screen "MTA-CompALTA" 1280x800, template "Plantilla"
   GraphicIOField "Plantilla_Campo ES gráfico_3" at 758,425 size 65x60
   GraphicIOField "Plantilla_Campo ES gráfico_4" at 685,353 size 65x60
   GraphicIOField "Plantilla_Campo ES gráfico_5" at 612,281 size 65x60
   GraphicIOField "Plantilla_Campo ES gráfico_2" at 539,209 size 65x60
   GraphicView "Visor de gráficos_2" at 492,46 size 254x172
   GraphicView "Visor de gráficos_18" at 492,46 size 254x172
   GraphicIOField "Plantilla_Campo ES gráfico_1" at 490,113 size 100x102
   GraphicView "Visor de gráficos_3" at 569,134 size 246x148
   ScreenModuleView "Faceplate_8_1" at 781,145 size 47x30
   GraphicView "Visor de gráficos_8" at 1175,577 size 29x50
   GraphicView "Visor de gráficos_7" at 885,605 size 391x113
   TextField "Plantilla_Campo de texto_1" at 1141,578 size 32x23
   IOField "Campo ES_1" at 943,632 size 108x28
   Button "Botón_7" at 1119,186 size 128x41
   Button "Botón_12" at 1119,234 size 128x41
   Button "Botón_13" at 1119,138 size 128x41
   Button "Botón_14" at 641,627 size 160x46
   TextField "Campo de texto_2" at 519,9 size 242x27
   ScreenModuleView "Faceplate_8_5" at 927,289 size 47x30
   ScreenModuleView "Faceplate_8_4" at 1000,361 size 47x30
   GraphicView "Visor de gráficos_19" at 569,134 size 246x148
   ScreenModuleView "Faceplate_8_2" at 854,217 size 47x30
   GraphicView "Visor de gráficos_4" at 642,206 size 246x148
   GraphicView "Visor de gráficos_22" at 642,206 size 246x148
   GraphicView "Visor de gráficos_5" at 715,278 size 246x148
   GraphicView "Visor de gráficos_21" at 715,278 size 246x148
   GraphicView "Visor de gráficos_6" at 788,350 size 246x148
   GraphicView "Visor de gráficos_20" at 788,350 size 246x148
   ScreenModuleView "Faceplate_8_3" at 1072,433 size 47x30
   ScreenModuleView "Faceplate_8_6" at 748,113 size 47x30
   Button "Botón_3" at 1181,68 size 48x46
   ScreenModuleView "Faceplate_8_7" at 1144,505 size 47x30
   GraphicIOField "Plantilla_Campo ES gráfico_6" at 831,497 size 65x60
   GraphicView "Visor de gráficos_1" at 861,422 size 246x148
   GraphicView "Visor de gráficos_9" at 861,422 size 246x148
   GraphicIOField "Campo ES gráfico_4" at 6,182 size 374x6
   SymbolicIOField "Campo ES simbólico_4" at 25,154 size 178x21
   TextField "Campo de texto_1" at 19,121 size 55x32
   GraphicIOField "Campo ES gráfico_5" at 118,341 size 374x6
   TextField "Campo de texto_6" at 127,280 size 67x32
   SymbolicIOField "Campo ES simbólico_5" at 137,313 size 186x21
   GraphicIOField "Campo ES gráfico_1" at 191,422 size 374x6
   TextField "Campo de texto_8" at 200,361 size 67x32
   SymbolicIOField "Campo ES simbólico_1" at 210,394 size 186x21
   GraphicIOField "Campo ES gráfico_3" at 44,262 size 373x6
   TextField "Campo de texto_10" at 53,201 size 67x32
   SymbolicIOField "Campo ES simbólico_3" at 63,234 size 194x21
   GraphicIOField "Campo ES gráfico_2" at 264,502 size 374x6
   TextField "Campo de texto_9" at 273,441 size 67x32
   SymbolicIOField "Campo ES simbólico_2" at 283,474 size 186x21
   GraphicIOField "Campo ES gráfico_16" at 337,582 size 374x6
   TextField "Campo de texto_3" at 346,521 size 67x32
   SymbolicIOField "Campo ES simbólico_11" at 356,554 size 186x21
   IOField "Campo ES_6" at 255,157 size 85x19
   IOField "Campo ES_2" at 367,316 size 85x19
   IOField "Campo ES_3" at 439,397 size 85x19
   IOField "Campo ES_5" at 292,237 size 85x19
   IOField "Campo ES_4" at 512,477 size 85x19
   IOField "Campo ES_7" at 585,557 size 85x19
   ScreenModuleView "Faceplate_6_1" at 283,125 size 57x28
   ScreenModuleView "Faceplate_6_5" at 395,284 size 57x28
   ScreenModuleView "Faceplate_6_4" at 468,365 size 57x28
   ScreenModuleView "Faceplate_6_2" at 321,205 size 57x28
   ScreenModuleView "Faceplate_6_3" at 541,445 size 57x28
   GraphicIOField "Campo ES gráfico_6" at 348,125 size 9x45
   GraphicIOField "Campo ES gráfico_9" at 357,125 size 9x45
   SymbolicIOField "Campo ES simbólico_6" at 86,124 size 160x29
   Button "Botón_11" at 6,116 size 374x64
   Switch "Interruptor_1" at 250,125 size 29x29
   Switch "Interruptor_10" at 863,114 size 40x40
   GraphicIOField "Campo ES gráfico_14" at 459,286 size 9x45
   GraphicIOField "Campo ES gráfico_15" at 468,286 size 9x45
   SymbolicIOField "Campo ES simbólico_10" at 195,283 size 160x29
   Button "Botón_6" at 118,275 size 374x64
   Switch "Interruptor_5" at 360,285 size 29x29
   Switch "Interruptor_9" at 1009,258 size 40x40
   GraphicIOField "Campo ES gráfico_12" at 532,367 size 9x45
   GraphicIOField "Campo ES gráfico_13" at 541,367 size 9x45
   Button "Botón_8" at 191,356 size 374x64
   SymbolicIOField "Campo ES simbólico_9" at 269,364 size 160x29
   Switch "Interruptor_4" at 433,366 size 29x29
   Switch "Interruptor_8" at 1082,330 size 40x40
   GraphicIOField "Campo ES gráfico_7" at 385,207 size 9x45
   GraphicIOField "Campo ES gráfico_10" at 394,207 size 9x45
   SymbolicIOField "Campo ES simbólico_7" at 120,204 size 160x29
   Switch "Interruptor_6" at 936,186 size 40x40
   GraphicIOField "Campo ES gráfico_8" at 605,447 size 9x45
   GraphicIOField "Campo ES gráfico_11" at 614,447 size 9x45
   SymbolicIOField "Campo ES simbólico_8" at 341,444 size 160x29
   Button "Botón_9" at 264,436 size 374x64
   Switch "Interruptor_3" at 504,445 size 29x29
   Switch "Interruptor_7" at 1155,402 size 40x40
   Switch "Interruptor_11" at 1228,474 size 40x40
   ScreenModuleView "Faceplate_6_6" at 614,525 size 57x28
   GraphicIOField "Campo ES gráfico_17" at 678,527 size 9x45
   GraphicIOField "Campo ES gráfico_18" at 687,527 size 9x45
   SymbolicIOField "Campo ES simbólico_12" at 414,524 size 160x29
   Button "Botón_1" at 337,516 size 374x64
   Switch "Interruptor_12" at 577,525 size 29x29
   Button "Botón_10" at 45,196 size 374x64
   Switch "Interruptor_2" at 284,206 size 29x29
   TextField "Campo de texto_4" at 591,208 size 309x29
   Button "Botón_2" at 912,202 size 128x41

screen "MTA-ALTAMC006" 1280x800, template "Plantilla-Alta-Cmp"
   Button "Botón_1" at 186,441 size 48x38
   Button "Botón_2" at 186,401 size 48x38
   Button "Botón_7" at 390,106 size 40x38
   Button "Botón_8" at 306,600 size 96x35
   TextField "Campo de texto_6" at 266,362 size 72x27
   TextField "Campo de texto_7" at 82,426 size 84x27
   TextField "Campo de texto_8" at 362,363 size 40x27
   TextField "Campo de texto_11" at 26,343 size 158x27
   GraphicIOField "Campo ES gráfico_3" at 294,402 size 16x78
   GraphicIOField "Campo ES gráfico_5" at 374,402 size 16x78
   SymbolicIOField "Campo ES simbólico_2" at 9,290 size 424x37
   TextField "Campo de texto_16" at 521,10 size 279x27
   TextField "Campo de texto_1" at 32,510 size 326x27
   TextField "Campo de texto_4" at 32,570 size 231x27
   TextField "Campo de texto_5" at 32,635 size 231x27
   Button "Botón_3" at 306,665 size 96x35
   GraphicIOField "Campo ES gráfico_2" at 10,280 size 422x6
   SymbolicIOField "Campo ES simbólico_4" at 19,246 size 290x21
   Button "Botón_6" at 13,154 size 88x62
   Switch "Interruptor_1" at 150,167 size 37x37
   ScreenModuleView "Faceplate_6_1" at 342,236 size 76x34
   ScreenModuleView "Faceplate_7_1" at 213,158 size 207x70
   IOField "Campo ES_7" at 20,535 size 173x35
   IOField "Campo ES_1" at 200,535 size 80x35
   IOField "Campo ES_2" at 20,595 size 173x35
   IOField "Campo ES_3" at 20,660 size 173x35

screen "EPROC-ALTAMS050" 1280x800, template "Plantilla-Alta-Sec"
   Button "Botón_3" at 467,294 size 40x38
   Button "Botón_4" at 411,540 size 96x35
   TextField "Campo de texto_6" at 37,450 size 326x27
   TextField "Campo de texto_4" at 37,510 size 201x27
   IOField "Campo ES_7" at 25,475 size 173x35
   IOField "Campo ES_1" at 205,475 size 80x35
   IOField "Campo ES_2" at 25,535 size 173x35
   GraphicIOField "Campo ES gráfico_3" at 21,434 size 511x6
   TextField "Campo de texto_3" at 46,356 size 89x39
   SymbolicIOField "Campo ES simbólico_3" at 48,392 size 242x21
   Switch "Interruptor_8" at 205,359 size 29x29
   ScreenModuleView "Faceplate_2_4" at 274,346 size 244x69

screen "EPROC-ALTAMS051" 1280x800, template "Plantilla-Alta-Sec"
   Button "Botón_3" at 467,294 size 40x38
   Button "Botón_4" at 411,540 size 96x35
   TextField "Campo de texto_6" at 37,450 size 326x27
   TextField "Campo de texto_4" at 37,510 size 201x27
   IOField "Campo ES_7" at 25,475 size 173x35
   IOField "Campo ES_1" at 205,475 size 80x35
   IOField "Campo ES_2" at 25,535 size 173x35
   GraphicIOField "Campo ES gráfico_9" at 21,434 size 511x6
   TextField "Campo de texto_1" at 46,356 size 89x39
   SymbolicIOField "Campo ES simbólico_9" at 48,392 size 242x21
   Switch "Interruptor_5" at 211,363 size 29x29
   ScreenModuleView "Faceplate_2_1" at 277,346 size 244x69

screen "EPROC-ALTAMS052" 1280x800, template "Plantilla-Alta-Sec"
   Button "Botón_3" at 467,294 size 40x38
   Button "Botón_4" at 411,540 size 96x35
   TextField "Campo de texto_6" at 37,450 size 326x27
   TextField "Campo de texto_4" at 37,510 size 201x27
   IOField "Campo ES_7" at 25,475 size 173x35
   IOField "Campo ES_1" at 205,475 size 80x35
   IOField "Campo ES_2" at 25,535 size 173x35
   GraphicIOField "Campo ES gráfico_1" at 21,434 size 511x6
   TextField "Campo de texto_1" at 46,356 size 89x39
   SymbolicIOField "Campo ES simbólico_1" at 48,392 size 242x21
   Switch "Interruptor_6" at 227,365 size 29x29
   ScreenModuleView "Faceplate_2_2" at 277,346 size 244x69

screen "EPROC-ALTAMS053" 1280x800, template "Plantilla-Alta-Sec"
   Button "Botón_3" at 467,294 size 40x38
   Button "Botón_4" at 411,540 size 96x35
   TextField "Campo de texto_6" at 37,450 size 326x27
   TextField "Campo de texto_4" at 37,510 size 201x27
   IOField "Campo ES_7" at 25,475 size 173x35
   IOField "Campo ES_1" at 205,475 size 80x35
   IOField "Campo ES_2" at 25,535 size 173x35
   IOField "Campo ES_6" at 351,413 size 85x19
   GraphicIOField "Campo ES gráfico_2" at 21,434 size 511x6
   TextField "Campo de texto_2" at 46,351 size 101x39
   SymbolicIOField "Campo ES simbólico_2" at 48,387 size 242x21
   Switch "Interruptor_7" at 227,360 size 29x29
   ScreenModuleView "Faceplate_2_3" at 276,346 size 244x69

screen "EPROC-BAJAMC060" 1280x800, template "Plantilla-Baja-Cmp"
   Button "Botón_4" at 1135,405 size 96x35
   TextField "Campo de texto_6" at 761,315 size 326x27
   TextField "Campo de texto_4" at 761,375 size 231x27
   Button "Botón_1" at 1135,470 size 96x35
   TextField "Campo de texto_1" at 761,440 size 231x27
   Button "Botón_2" at 1135,535 size 96x35
   TextField "Campo de texto_2" at 761,505 size 231x27
   Button "Botón_3" at 1135,600 size 96x35
   TextField "Campo de texto_3" at 761,570 size 231x27
   Button "Botón_5" at 1135,665 size 96x35
   TextField "Campo de texto_7" at 761,635 size 231x27
   Button "Botón_6" at 1199,168 size 40x38
   GraphicIOField "Campo ES gráfico_4" at 746,294 size 511x6
   TextField "Campo de texto_5" at 771,224 size 116x39
   SymbolicIOField "Campo ES simbólico_9" at 773,260 size 242x21
   Switch "Interruptor_5" at 1108,242 size 91x31
   IOField "Campo ES_7" at 749,340 size 173x35
   IOField "Campo ES_1" at 929,340 size 80x35
   IOField "Campo ES_2" at 749,400 size 173x35
   IOField "Campo ES_3" at 749,465 size 173x35
   IOField "Campo ES_4" at 749,530 size 173x35
   IOField "Campo ES_5" at 749,595 size 173x35
   IOField "Campo ES_6" at 749,660 size 173x35

screen "EPROC-BAJAMC061" 1280x800, template "Plantilla-Baja-Cmp"
   Button "Botón_4" at 1135,405 size 96x35
   TextField "Campo de texto_6" at 761,315 size 326x27
   TextField "Campo de texto_4" at 761,375 size 231x27
   Button "Botón_1" at 1135,470 size 96x35
   TextField "Campo de texto_1" at 761,440 size 231x27
   Button "Botón_2" at 1135,535 size 96x35
   TextField "Campo de texto_2" at 761,505 size 231x27
   Button "Botón_3" at 1135,600 size 96x35
   TextField "Campo de texto_3" at 761,570 size 231x27
   Button "Botón_5" at 1135,665 size 96x35
   TextField "Campo de texto_7" at 761,635 size 231x27
   Button "Botón_6" at 1199,168 size 40x38
   IOField "Campo ES_7" at 749,340 size 173x35
   IOField "Campo ES_1" at 929,340 size 80x35
   IOField "Campo ES_2" at 749,400 size 173x35
   IOField "Campo ES_3" at 749,465 size 173x35
   IOField "Campo ES_4" at 749,530 size 173x35
   IOField "Campo ES_5" at 749,595 size 173x35
   IOField "Campo ES_6" at 749,660 size 173x35
   GraphicIOField "Campo ES gráfico_3" at 746,293 size 510x6
   TextField "Campo de texto_5" at 771,224 size 116x39
   SymbolicIOField "Campo ES simbólico_8" at 773,260 size 242x21
   Switch "Interruptor_4" at 974,228 size 29x29
   ScreenModuleView "Faceplate_1_1" at 1018,228 size 236x58

screen "EPROC-BAJAMC062" 1280x800, template "Plantilla-Baja-Cmp"
   Button "Botón_4" at 1135,405 size 96x35
   TextField "Campo de texto_6" at 761,315 size 326x27
   TextField "Campo de texto_4" at 761,375 size 231x27
   Button "Botón_1" at 1135,470 size 96x35
   TextField "Campo de texto_1" at 761,440 size 231x27
   Button "Botón_2" at 1135,535 size 96x35
   TextField "Campo de texto_2" at 761,505 size 231x27
   Button "Botón_3" at 1135,600 size 96x35
   TextField "Campo de texto_3" at 761,570 size 231x27
   Button "Botón_5" at 1135,665 size 96x35
   TextField "Campo de texto_7" at 761,635 size 231x27
   Button "Botón_6" at 1199,168 size 40x38
   IOField "Campo ES_7" at 749,340 size 173x35
   IOField "Campo ES_1" at 929,340 size 80x35
   IOField "Campo ES_2" at 749,400 size 173x35
   IOField "Campo ES_3" at 749,465 size 173x35
   IOField "Campo ES_4" at 749,530 size 173x35
   IOField "Campo ES_5" at 749,595 size 173x35
   IOField "Campo ES_6" at 749,660 size 173x35
   GraphicIOField "Campo ES gráfico_2" at 747,293 size 507x6
   TextField "Campo de texto_5" at 771,224 size 116x39
   SymbolicIOField "Campo ES simbólico_7" at 773,260 size 242x21
   Switch "Interruptor_3" at 970,227 size 29x29
   ScreenModuleView "Faceplate_1_3" at 1013,227 size 236x58

screen "EPROC-BAJAMC063" 1280x800, template "Plantilla-Baja-Cmp"
   Button "Botón_4" at 1135,405 size 96x35
   TextField "Campo de texto_6" at 761,315 size 326x27
   TextField "Campo de texto_4" at 761,375 size 231x27
   Button "Botón_1" at 1135,470 size 96x35
   TextField "Campo de texto_1" at 761,440 size 231x27
   Button "Botón_2" at 1135,535 size 96x35
   TextField "Campo de texto_2" at 761,505 size 231x27
   Button "Botón_3" at 1135,600 size 96x35
   TextField "Campo de texto_3" at 761,570 size 231x27
   Button "Botón_5" at 1135,665 size 96x35
   TextField "Campo de texto_7" at 761,635 size 231x27
   Button "Botón_6" at 1199,168 size 40x38
   IOField "Campo ES_7" at 749,340 size 173x35
   IOField "Campo ES_1" at 929,340 size 80x35
   IOField "Campo ES_2" at 749,400 size 173x35
   IOField "Campo ES_3" at 749,465 size 173x35
   IOField "Campo ES_4" at 749,530 size 173x35
   IOField "Campo ES_5" at 749,595 size 173x35
   IOField "Campo ES_6" at 749,660 size 173x35
   GraphicIOField "Campo ES gráfico_1" at 746,293 size 507x6
   TextField "Campo de texto_8" at 763,224 size 91x39
   SymbolicIOField "Campo ES simbólico_6" at 765,260 size 242x21
   Switch "Interruptor_2" at 967,227 size 29x29
   ScreenModuleView "Faceplate_1_4" at 1014,226 size 236x58

screen "EPROC-BAJAMC064" 1280x800, template "Plantilla-Baja-Cmp"
   Button "Botón_4" at 1135,405 size 96x35
   TextField "Campo de texto_6" at 761,315 size 326x27
   TextField "Campo de texto_4" at 761,375 size 231x27
   Button "Botón_1" at 1135,470 size 96x35
   TextField "Campo de texto_1" at 761,440 size 231x27
   Button "Botón_2" at 1135,535 size 96x35
   TextField "Campo de texto_2" at 761,505 size 231x27
   Button "Botón_3" at 1135,600 size 96x35
   TextField "Campo de texto_3" at 761,570 size 231x27
   Button "Botón_5" at 1135,665 size 96x35
   TextField "Campo de texto_7" at 761,635 size 231x27
   Button "Botón_6" at 1199,168 size 40x38
   IOField "Campo ES_7" at 749,340 size 173x35
   IOField "Campo ES_1" at 929,340 size 80x35
   IOField "Campo ES_2" at 749,400 size 173x35
   IOField "Campo ES_3" at 749,465 size 173x35
   IOField "Campo ES_4" at 749,530 size 173x35
   IOField "Campo ES_5" at 749,595 size 173x35
   IOField "Campo ES_6" at 749,660 size 173x35
   GraphicIOField "Campo ES gráfico_5" at 747,294 size 507x6
   TextField "Campo de texto_9" at 771,224 size 100x39
   SymbolicIOField "Campo ES simbólico_5" at 773,260 size 242x21
   Switch "Interruptor_1" at 969,227 size 29x29
   ScreenModuleView "Faceplate_1_5" at 1016,227 size 236x58

screen "EPROC-BAJAMS054" 1280x800, template "Plantilla-Baja-Sec"
   TextField "Campo de texto_1" at 758,509 size 326x27
   Button "Botón_4" at 1032,599 size 96x35
   TextField "Campo de texto_4" at 758,569 size 231x27
   TextField "Campo de texto_5" at 758,634 size 231x27
   Button "Botón_5" at 1032,664 size 96x35
   Button "Botón_6" at 1188,358 size 40x38
   IOField "Campo ES_7" at 746,534 size 173x35
   IOField "Campo ES_1" at 926,534 size 80x35
   IOField "Campo ES_2" at 746,594 size 173x35
   IOField "Campo ES_3" at 746,659 size 173x35
   GraphicIOField "Campo ES gráfico_3" at 736,489 size 510x6
   TextField "Campo de texto_6" at 761,411 size 116x39
   SymbolicIOField "Campo ES simbólico_8" at 763,447 size 242x21
   ScreenModuleView "Faceplate_3_1" at 1015,411 size 213x73

screen "EPROC-BAJAMS055" 1280x800, template "Plantilla-Baja-Sec"
   TextField "Campo de texto_1" at 758,509 size 326x27
   Button "Botón_4" at 1032,599 size 96x35
   TextField "Campo de texto_4" at 758,569 size 231x27
   TextField "Campo de texto_5" at 758,634 size 231x27
   Button "Botón_5" at 1032,664 size 96x35
   Button "Botón_6" at 1188,358 size 40x38
   IOField "Campo ES_7" at 746,534 size 173x35
   IOField "Campo ES_1" at 926,534 size 80x35
   IOField "Campo ES_2" at 746,594 size 173x35
   IOField "Campo ES_3" at 746,659 size 173x35
   GraphicIOField "Campo ES gráfico_4" at 736,489 size 511x6
   TextField "Campo de texto_2" at 761,411 size 116x39
   SymbolicIOField "Campo ES simbólico_9" at 763,447 size 242x21
   ScreenModuleView "Faceplate_3_2" at 1020,411 size 213x73

screen "Imagen_1" 1280x800
   GraphicIOField "Campo ES gráfico_3" at 736,489 size 510x6
   TextField "Campo de texto_6" at 761,411 size 116x39
   SymbolicIOField "Campo ES simbólico_8" at 763,447 size 242x21
   ScreenModuleView "Faceplate_3_1" at 1015,411 size 213x73

Template "Plantilla" 1280x800
   Button "Plantilla_6" at 1196,741 size 81x58
   Button "Plantilla_1" at 1037,749 size 78x50
   Button "Plantilla_3" at 717,748 size 78x50
   Button "Plantilla_4" at 877,748 size 78x50
   Button "Plantilla_5" at 957,748 size 78x50
   Button "Plantilla_7" at 479,748 size 78x50
   Button "Plantilla_8" at 161,748 size 78x50
   Button "Plantilla_9" at 81,748 size 78x50
   Button "Plantilla_10" at 1117,741 size 78x58
   Button "Plantilla_12" at 638,748 size 78x50
   Button "Plantilla_13" at 400,748 size 78x50
   Button "Plantilla_14" at 321,748 size 78x50
   Button "Plantilla_15" at 558,748 size 78x50
   Button "Plantilla_16" at 241,748 size 78x50
   Button "Plantilla_17" at 1,740 size 78x58
   GraphicView "Plantilla_Visor de gráficos_1" at 80,740 size 78x6
   GraphicView "Plantilla_Visor de gráficos_2" at 160,740 size 78x6
   GraphicView "Plantilla_Visor de gráficos_3" at 478,740 size 78x6
   GraphicView "Plantilla_Visor de gráficos_4" at 240,740 size 78x6
   GraphicView "Plantilla_Visor de gráficos_5" at 557,740 size 78x6
   GraphicView "Plantilla_Visor de gráficos_6" at 320,740 size 78x6
   GraphicView "Plantilla_Visor de gráficos_7" at 399,740 size 78x6
   GraphicView "Plantilla_Visor de gráficos_11" at 637,740 size 78x6
   GraphicView "Plantilla_Visor de gráficos_8" at 80,740 size 78x6
   GraphicView "Plantilla_Visor de gráficos_9" at 160,740 size 78x6
   GraphicView "Plantilla_Visor de gráficos_10" at 478,740 size 78x6
   GraphicView "Plantilla_Visor de gráficos_12" at 240,740 size 78x6
   GraphicView "Plantilla_Visor de gráficos_13" at 557,740 size 78x6
   GraphicView "Plantilla_Visor de gráficos_14" at 320,740 size 78x6
   GraphicView "Plantilla_Visor de gráficos_15" at 399,740 size 78x6
   GraphicView "Plantilla_Visor de gráficos_16" at 637,740 size 78x6
   TextField "Plantilla_Campo de texto_2" at 521,711 size 69x18
   TextField "Plantilla_Campo de texto_4" at 323,711 size 68x18
   TextField "Plantilla_Campo de texto_1" at 139,711 size 40x18
   Button "Plantilla_11" at 797,748 size 78x50
   GraphicView "Plantilla_Visor de gráficos_18" at 717,740 size 78x6
   GraphicView "Plantilla_Visor de gráficos_19" at 797,740 size 78x6
   GraphicView "Plantilla_Visor de gráficos_20" at 877,740 size 78x6
   GraphicView "Plantilla_Visor de gráficos_21" at 957,740 size 78x6
   GraphicView "Plantilla_Visor de gráficos_22" at 1037,741 size 78x6
   GraphicView "Plantilla_Visor de gráficos_23" at 1037,741 size 78x6
   GraphicView "Plantilla_Visor de gráficos_24" at 877,740 size 78x6
   Group "Group" at 1,716 size 1276x83
   GraphicView "Plantilla_Visor de gráficos_26" at 68,9 size 91x26
   GraphicView "Plantilla_Visor de gráficos_27" at 9,8 size 49x29
   TextField "Plantilla_Campo de texto_3" at 32,732 size 696x50
   Button "Plantilla_Botón_1" at 1232,724 size 37x34
   Button "Plantilla_Botón_2" at 945,735 size 112x46
   Button "Plantilla_Botón_3" at 1065,735 size 112x46

Template "Plantilla-Alta-Cmp" 1280x800
   TextField "Plantilla_Campo de texto_5" at 32,731 size 696x50
   Button "Plantilla_Botón_1" at 1232,723 size 37x34
   Button "Plantilla_Botón_2" at 945,734 size 112x46
   Button "Plantilla_Botón_3" at 1065,734 size 112x46
   GraphicView "Visor de gráficos_8" at 1175,577 size 29x50
   GraphicView "Visor de gráficos_7" at 885,605 size 391x113
   Button "Plantilla_6" at 1196,741 size 81x58
   GraphicView "Plantilla_Visor de gráficos_17" at 4,4 size 87x38
   Button "Plantilla_7" at 479,748 size 78x50
   Button "Plantilla_8" at 161,748 size 78x50
   Button "Plantilla_9" at 81,748 size 78x50
   Button "Plantilla_12" at 638,748 size 78x50
   Button "Plantilla_13" at 400,748 size 78x50
   Button "Plantilla_14" at 321,748 size 78x50
   Button "Plantilla_15" at 558,748 size 78x50
   Button "Plantilla_16" at 241,748 size 78x50
   Button "Plantilla_17" at 1,740 size 78x58
   GraphicView "Plantilla_Visor de gráficos_1" at 80,740 size 78x6
   GraphicView "Plantilla_Visor de gráficos_2" at 160,740 size 78x6
   GraphicView "Plantilla_Visor de gráficos_3" at 478,740 size 78x6
   GraphicView "Plantilla_Visor de gráficos_4" at 240,740 size 78x6
   GraphicView "Plantilla_Visor de gráficos_5" at 557,740 size 78x6
   GraphicView "Plantilla_Visor de gráficos_6" at 320,740 size 78x6
   GraphicView "Plantilla_Visor de gráficos_7" at 399,740 size 78x6
   GraphicView "Plantilla_Visor de gráficos_11" at 637,740 size 78x6
   GraphicView "Plantilla_Visor de gráficos_8" at 80,740 size 78x6
   GraphicView "Plantilla_Visor de gráficos_9" at 160,740 size 78x6
   GraphicView "Plantilla_Visor de gráficos_10" at 478,740 size 78x6
   GraphicView "Plantilla_Visor de gráficos_12" at 240,740 size 78x6
   GraphicView "Plantilla_Visor de gráficos_13" at 557,740 size 78x6
   GraphicView "Plantilla_Visor de gráficos_14" at 320,740 size 78x6
   GraphicView "Plantilla_Visor de gráficos_15" at 399,740 size 78x6
   GraphicView "Plantilla_Visor de gráficos_16" at 637,740 size 78x6
   TextField "Plantilla_Campo de texto_2" at 521,711 size 69x18
   TextField "Plantilla_Campo de texto_4" at 323,711 size 68x18
   TextField "Plantilla_Campo de texto_3" at 139,711 size 40x18
   Button "Plantilla_3" at 717,748 size 78x50
   Button "Plantilla_5" at 957,748 size 78x50
   Button "Plantilla_11" at 797,748 size 78x50
   GraphicView "Plantilla_Visor de gráficos_18" at 717,740 size 78x6
   GraphicView "Plantilla_Visor de gráficos_19" at 797,740 size 78x6
   GraphicView "Plantilla_Visor de gráficos_20" at 877,740 size 78x6
   GraphicView "Plantilla_Visor de gráficos_21" at 957,740 size 78x6
   GraphicView "Plantilla_Visor de gráficos_22" at 1037,740 size 78x6
   GraphicView "Plantilla_Visor de gráficos_23" at 1037,740 size 78x6
   Button "Plantilla_1" at 1037,749 size 78x50
   Button "Plantilla_2" at 1117,741 size 78x58
   Button "Plantilla_4" at 877,748 size 78x50
   GraphicView "Plantilla_Visor de gráficos_24" at 877,740 size 78x6
   GraphicView "Plantilla_Visor de gráficos_25" at 877,740 size 78x6
   Group "Group" at 1,715 size 1276x84
   GraphicView "Plantilla_Visor de gráficos_26" at 68,9 size 91x26
   GraphicView "Plantilla_Visor de gráficos_27" at 9,8 size 49x29
   GraphicView "Visor de gráficos_2" at 492,46 size 254x172
   GraphicIOField "Plantilla_Campo ES gráfico_3" at 758,425 size 65x60
   GraphicIOField "Plantilla_Campo ES gráfico_4" at 685,353 size 65x60
   GraphicIOField "Plantilla_Campo ES gráfico_5" at 612,281 size 65x60
   GraphicIOField "Plantilla_Campo ES gráfico_2" at 539,209 size 65x60
   GraphicView "Visor de gráficos_18" at 492,46 size 254x172
   GraphicIOField "Plantilla_Campo ES gráfico_1" at 490,113 size 100x102
   GraphicView "Visor de gráficos_3" at 569,134 size 246x148
   ScreenModuleView "Faceplate_8_1" at 781,145 size 47x30
   TextField "Plantilla_Campo de texto_1" at 1141,578 size 35x23
   IOField "Campo ES_1" at 943,632 size 108x28
   Button "Botón_7" at 1119,186 size 128x41
   Button "Botón_12" at 1119,234 size 128x41
   Button "Botón_13" at 1119,138 size 128x41
   ScreenModuleView "Faceplate_8_5" at 927,289 size 47x30
   ScreenModuleView "Faceplate_8_4" at 1000,361 size 47x30
   GraphicView "Visor de gráficos_19" at 569,134 size 246x148
   ScreenModuleView "Faceplate_8_2" at 854,217 size 47x30
   GraphicView "Visor de gráficos_4" at 642,206 size 246x148
   GraphicView "Visor de gráficos_22" at 642,206 size 246x148
   GraphicView "Visor de gráficos_5" at 715,278 size 246x148
   GraphicView "Visor de gráficos_21" at 715,278 size 246x148
   GraphicView "Visor de gráficos_6" at 788,350 size 246x148
   GraphicView "Visor de gráficos_20" at 788,350 size 246x148
   ScreenModuleView "Faceplate_8_3" at 1072,433 size 47x30
   ScreenModuleView "Faceplate_8_6" at 748,113 size 47x30
   ScreenModuleView "Faceplate_8_7" at 1144,505 size 47x30
   GraphicIOField "Plantilla_Campo ES gráfico_6" at 831,497 size 65x60
   GraphicView "Visor de gráficos_1" at 861,422 size 246x148
   GraphicView "Visor de gráficos_9" at 861,422 size 246x148
   Switch "Interruptor_10" at 863,114 size 40x40
   Switch "Interruptor_9" at 1009,258 size 40x40
   Switch "Interruptor_8" at 1082,330 size 40x40
   Switch "Interruptor_6" at 936,186 size 40x40
   Switch "Interruptor_7" at 1155,402 size 40x40
   Switch "Interruptor_11" at 1228,474 size 40x40

Template "Plantilla-Alta-Sec" 1280x800
   Button "Plantilla_6" at 1196,741 size 81x58
   GraphicView "Plantilla_Visor de gráficos_17" at 4,4 size 87x38
   Button "Plantilla_7" at 479,748 size 78x50
   Button "Plantilla_8" at 161,748 size 78x50
   Button "Plantilla_9" at 81,748 size 78x50
   Button "Plantilla_12" at 638,748 size 78x50
   Button "Plantilla_13" at 400,748 size 78x50
   Button "Plantilla_14" at 321,748 size 78x50
   Button "Plantilla_15" at 558,748 size 78x50
   Button "Plantilla_16" at 241,748 size 78x50
   Button "Plantilla_17" at 1,740 size 78x58
   GraphicView "Plantilla_Visor de gráficos_1" at 80,740 size 78x6
   GraphicView "Plantilla_Visor de gráficos_2" at 160,740 size 78x6
   GraphicView "Plantilla_Visor de gráficos_3" at 478,740 size 78x6
   GraphicView "Plantilla_Visor de gráficos_4" at 240,740 size 78x6
   GraphicView "Plantilla_Visor de gráficos_5" at 557,740 size 78x6
   GraphicView "Plantilla_Visor de gráficos_6" at 320,740 size 78x6
   GraphicView "Plantilla_Visor de gráficos_7" at 399,740 size 78x6
   GraphicView "Plantilla_Visor de gráficos_11" at 637,740 size 78x6
   GraphicView "Plantilla_Visor de gráficos_8" at 80,740 size 78x6
   GraphicView "Plantilla_Visor de gráficos_9" at 160,740 size 78x6
   GraphicView "Plantilla_Visor de gráficos_10" at 478,740 size 78x6
   GraphicView "Plantilla_Visor de gráficos_12" at 240,740 size 78x6
   GraphicView "Plantilla_Visor de gráficos_13" at 557,740 size 78x6
   GraphicView "Plantilla_Visor de gráficos_14" at 320,740 size 78x6
   GraphicView "Plantilla_Visor de gráficos_15" at 399,740 size 78x6
   GraphicView "Plantilla_Visor de gráficos_16" at 637,740 size 78x6
   TextField "Plantilla_Campo de texto_2" at 521,711 size 69x18
   TextField "Plantilla_Campo de texto_4" at 323,711 size 68x18
   TextField "Plantilla_Campo de texto_3" at 139,711 size 40x18
   Button "Plantilla_3" at 717,748 size 78x50
   Button "Plantilla_5" at 957,748 size 78x50
   Button "Plantilla_11" at 797,748 size 78x50
   GraphicView "Plantilla_Visor de gráficos_18" at 717,740 size 78x6
   GraphicView "Plantilla_Visor de gráficos_19" at 797,740 size 78x6
   GraphicView "Plantilla_Visor de gráficos_20" at 877,740 size 78x6
   GraphicView "Plantilla_Visor de gráficos_21" at 957,740 size 78x6
   GraphicView "Plantilla_Visor de gráficos_22" at 1037,740 size 78x6
   GraphicView "Plantilla_Visor de gráficos_23" at 1037,740 size 78x6
   Button "Plantilla_1" at 1037,749 size 78x50
   Button "Plantilla_2" at 1117,741 size 78x58
   Button "Plantilla_4" at 877,748 size 78x50
   GraphicView "Plantilla_Visor de gráficos_24" at 877,740 size 78x6
   GraphicView "Plantilla_Visor de gráficos_25" at 877,740 size 78x6
   Group "Group" at 1,715 size 1276x84
   GraphicView "Plantilla_Visor de gráficos_26" at 68,9 size 91x26
   GraphicView "Plantilla_Visor de gráficos_27" at 9,8 size 49x29
   GraphicIOField "Campo ES gráfico_4" at 981,258 size 280x222
   GraphicView "Visor de gráficos_4" at 999,137 size 234x314
   GraphicView "Visor de gráficos_15" at 999,137 size 234x314
   GraphicIOField "Campo ES gráfico_8" at 571,212 size 366x99
   GraphicView "Visor de gráficos_3" at 592,100 size 363x184
   GraphicView "Visor de gráficos_5" at 592,100 size 363x184
   GraphicIOField "Campo ES gráfico_7" at 674,357 size 309x81
   GraphicView "Visor de gráficos_2" at 696,255 size 292x158
   GraphicView "Visor de gráficos_6" at 695,255 size 294x158
   GraphicIOField "Campo ES gráfico_6" at 765,490 size 338x86
   GraphicView "Visor de gráficos_1" at 786,405 size 292x142
   GraphicView "Visor de gráficos_14" at 786,405 size 292x142
   TextField "Plantilla_Campo de texto_5" at 32,731 size 696x50
   Button "Plantilla_Botón_1" at 1232,723 size 37x34
   Button "Plantilla_Botón_2" at 945,734 size 112x46
   Button "Plantilla_Botón_3" at 1065,734 size 112x46
   Switch "Interruptor_1" at 640,315 size 40x40
   Switch "Interruptor_2" at 731,440 size 40x40
   Switch "Interruptor_3" at 540,176 size 40x40
   Switch "Interruptor_4" at 1212,488 size 40x40

Template "Plantilla-Baja-Cmp" 1280x800
   Button "Plantilla_6" at 1196,741 size 81x58
   GraphicView "Plantilla_Visor de gráficos_17" at 4,4 size 87x38
   Button "Plantilla_7" at 479,748 size 78x50
   Button "Plantilla_8" at 161,748 size 78x50
   Button "Plantilla_9" at 81,748 size 78x50
   Button "Plantilla_12" at 638,748 size 78x50
   Button "Plantilla_13" at 400,748 size 78x50
   Button "Plantilla_14" at 321,748 size 78x50
   Button "Plantilla_15" at 558,748 size 78x50
   Button "Plantilla_16" at 241,748 size 78x50
   Button "Plantilla_17" at 1,740 size 78x58
   GraphicView "Plantilla_Visor de gráficos_1" at 80,740 size 78x6
   GraphicView "Plantilla_Visor de gráficos_2" at 160,740 size 78x6
   GraphicView "Plantilla_Visor de gráficos_3" at 478,740 size 78x6
   GraphicView "Plantilla_Visor de gráficos_4" at 240,740 size 78x6
   GraphicView "Plantilla_Visor de gráficos_5" at 557,740 size 78x6
   GraphicView "Plantilla_Visor de gráficos_6" at 320,740 size 78x6
   GraphicView "Plantilla_Visor de gráficos_7" at 399,740 size 78x6
   GraphicView "Plantilla_Visor de gráficos_11" at 637,740 size 78x6
   GraphicView "Plantilla_Visor de gráficos_8" at 80,740 size 78x6
   GraphicView "Plantilla_Visor de gráficos_9" at 160,740 size 78x6
   GraphicView "Plantilla_Visor de gráficos_10" at 478,740 size 78x6
   GraphicView "Plantilla_Visor de gráficos_12" at 240,740 size 78x6
   GraphicView "Plantilla_Visor de gráficos_13" at 557,740 size 78x6
   GraphicView "Plantilla_Visor de gráficos_14" at 320,740 size 78x6
   GraphicView "Plantilla_Visor de gráficos_15" at 399,740 size 78x6
   GraphicView "Plantilla_Visor de gráficos_16" at 637,740 size 78x6
   TextField "Plantilla_Campo de texto_2" at 521,711 size 69x18
   TextField "Plantilla_Campo de texto_4" at 323,711 size 68x18
   TextField "Plantilla_Campo de texto_3" at 139,711 size 40x18
   Button "Plantilla_3" at 717,748 size 78x50
   Button "Plantilla_5" at 957,748 size 78x50
   Button "Plantilla_11" at 797,748 size 78x50
   GraphicView "Plantilla_Visor de gráficos_18" at 717,740 size 78x6
   GraphicView "Plantilla_Visor de gráficos_19" at 797,740 size 78x6
   GraphicView "Plantilla_Visor de gráficos_20" at 877,740 size 78x6
   GraphicView "Plantilla_Visor de gráficos_21" at 957,740 size 78x6
   GraphicView "Plantilla_Visor de gráficos_22" at 1037,740 size 78x6
   GraphicView "Plantilla_Visor de gráficos_23" at 1037,740 size 78x6
   Button "Plantilla_1" at 1037,749 size 78x50
   Button "Plantilla_2" at 1117,741 size 78x58
   Button "Plantilla_4" at 877,748 size 78x50
   GraphicView "Plantilla_Visor de gráficos_24" at 877,740 size 78x6
   GraphicView "Plantilla_Visor de gráficos_25" at 877,740 size 78x6
   Group "Group" at 1,715 size 1276x84
   GraphicView "Plantilla_Visor de gráficos_26" at 68,9 size 91x26
   GraphicView "Plantilla_Visor de gráficos_27" at 9,8 size 49x29
   GraphicIOField "Campo ES gráfico_10" at 491,153 size 189x58
   GraphicIOField "Campo ES gráfico_9" at 427,241 size 189x58
   GraphicIOField "Campo ES gráfico_7" at 387,316 size 178x52
   GraphicIOField "Campo ES gráfico_6" at 340,387 size 178x52
   GraphicIOField "Campo ES gráfico_8" at 275,454 size 197x58
   GraphicView "Visor de gráficos_1" at 467,72 size 269x127
   GraphicView "Visor de gráficos_7" at 467,72 size 269x127
   GraphicView "Visor de gráficos_2" at 403,160 size 269x127
   GraphicView "Visor de gráficos_8" at 403,160 size 269x127
   GraphicView "Visor de gráficos_3" at 315,232 size 269x127
   GraphicView "Visor de gráficos_9" at 315,232 size 269x127
   GraphicView "Visor de gráficos_4" at 267,304 size 269x127
   GraphicView "Visor de gráficos_10" at 267,304 size 269x127
   GraphicView "Visor de gráficos_5" at 243,376 size 213x127
   GraphicView "Visor de gráficos_11" at 243,376 size 213x127
   GraphicView "Visor de gráficos_6" at 132,415 size 202x177
   IOField "Campo ES_1" at 161,449 size 148x28
   GraphicView "Visor de gráficos_12" at 18,528 size 229x141
   GraphicIOField "Campo ES gráfico_11" at 68,583 size 48x46
   GraphicIOField "Campo ES gráfico_12" at 160,500 size 17x32
   GraphicIOField "Campo ES gráfico_13" at 40,563 size 169x87
   GraphicView "Visor de gráficos_18" at 440,520 size 40x40
   GraphicView "Visor de gráficos_19" at 440,520 size 40x40
   Button "Botón_11" at 440,520 size 40x40
   GraphicView "Visor de gráficos_17" at 226,528 size 229x141
   GraphicIOField "Campo ES gráfico_15" at 286,586 size 48x47
   GraphicIOField "Campo ES gráfico_16" at 368,500 size 18x34
   GraphicIOField "Campo ES gráfico_17" at 261,565 size 156x84
   GraphicView "Visor de gráficos_13" at 37,520 size 40x40
   GraphicView "Visor de gráficos_14" at 37,520 size 40x40
   Button "Botón_6" at 37,520 size 40x40
   TextField "Campo de texto_4" at 48,674 size 122x19
   TextField "Campo de texto_10" at 251,674 size 122x19
   TextField "Plantilla_Campo de texto_5" at 32,731 size 696x50
   Button "Plantilla_Botón_1" at 1232,723 size 37x34
   Button "Plantilla_Botón_2" at 945,734 size 112x46
   Button "Plantilla_Botón_3" at 1065,734 size 112x46
   Switch "Interruptor_6" at 313,243 size 40x40
   Switch "Interruptor_7" at 265,323 size 40x40
   Switch "Interruptor_9" at 365,171 size 40x40
   Switch "Interruptor_10" at 429,83 size 40x40

Template "Plantilla-Baja-Sec" 1280x800
   Button "Plantilla_6" at 1196,741 size 81x58
   GraphicView "Plantilla_Visor de gráficos_17" at 4,4 size 87x38
   Button "Plantilla_7" at 479,748 size 78x50
   Button "Plantilla_8" at 161,748 size 78x50
   Button "Plantilla_9" at 81,748 size 78x50
   Button "Plantilla_12" at 638,748 size 78x50
   Button "Plantilla_13" at 400,748 size 78x50
   Button "Plantilla_14" at 321,748 size 78x50
   Button "Plantilla_15" at 558,748 size 78x50
   Button "Plantilla_16" at 241,748 size 78x50
   Button "Plantilla_17" at 1,740 size 78x58
   GraphicView "Plantilla_Visor de gráficos_1" at 80,740 size 78x6
   GraphicView "Plantilla_Visor de gráficos_2" at 160,740 size 78x6
   GraphicView "Plantilla_Visor de gráficos_3" at 478,740 size 78x6
   GraphicView "Plantilla_Visor de gráficos_4" at 240,740 size 78x6
   GraphicView "Plantilla_Visor de gráficos_5" at 557,740 size 78x6
   GraphicView "Plantilla_Visor de gráficos_6" at 320,740 size 78x6
   GraphicView "Plantilla_Visor de gráficos_7" at 399,740 size 78x6
   GraphicView "Plantilla_Visor de gráficos_11" at 637,740 size 78x6
   GraphicView "Plantilla_Visor de gráficos_8" at 80,740 size 78x6
   GraphicView "Plantilla_Visor de gráficos_9" at 160,740 size 78x6
   GraphicView "Plantilla_Visor de gráficos_10" at 478,740 size 78x6
   GraphicView "Plantilla_Visor de gráficos_12" at 240,740 size 78x6
   GraphicView "Plantilla_Visor de gráficos_13" at 557,740 size 78x6
   GraphicView "Plantilla_Visor de gráficos_14" at 320,740 size 78x6
   GraphicView "Plantilla_Visor de gráficos_15" at 399,740 size 78x6
   GraphicView "Plantilla_Visor de gráficos_16" at 637,740 size 78x6
   TextField "Plantilla_Campo de texto_2" at 521,711 size 69x18
   TextField "Plantilla_Campo de texto_4" at 323,711 size 68x18
   TextField "Plantilla_Campo de texto_3" at 139,711 size 40x18
   Button "Plantilla_3" at 717,748 size 78x50
   Button "Plantilla_5" at 957,748 size 78x50
   Button "Plantilla_11" at 797,748 size 78x50
   GraphicView "Plantilla_Visor de gráficos_18" at 717,740 size 78x6
   GraphicView "Plantilla_Visor de gráficos_19" at 797,740 size 78x6
   GraphicView "Plantilla_Visor de gráficos_20" at 877,740 size 78x6
   GraphicView "Plantilla_Visor de gráficos_21" at 957,740 size 78x6
   GraphicView "Plantilla_Visor de gráficos_22" at 1037,740 size 78x6
   GraphicView "Plantilla_Visor de gráficos_23" at 1037,740 size 78x6
   Button "Plantilla_1" at 1037,749 size 78x50
   Button "Plantilla_2" at 1117,741 size 78x58
   Button "Plantilla_4" at 877,748 size 78x50
   GraphicView "Plantilla_Visor de gráficos_24" at 877,740 size 78x6
   GraphicView "Plantilla_Visor de gráficos_25" at 877,740 size 78x6
   Group "Group" at 1,715 size 1276x84
   GraphicView "Plantilla_Visor de gráficos_26" at 68,9 size 91x26
   GraphicView "Plantilla_Visor de gráficos_27" at 9,8 size 49x29
   GraphicIOField "Campo ES gráfico_1" at 289,314 size 285x90
   GraphicView "Visor de gráficos_2" at 333,200 size 201x179
   GraphicIOField "Campo ES gráfico_8" at 159,455 size 269x90
   GraphicView "Visor de gráficos_4" at 333,200 size 201x179
   GraphicView "Visor de gráficos_1" at 192,341 size 201x179
   GraphicView "Visor de gráficos_3" at 192,341 size 201x179
   TextField "Plantilla_Campo de texto_5" at 32,731 size 696x50
   Button "Plantilla_Botón_1" at 1232,723 size 37x34
   Button "Plantilla_Botón_2" at 945,734 size 112x46
   Button "Plantilla_Botón_3" at 1065,734 size 112x46
   Switch "Interruptor_7" at 271,262 size 40x40
   Switch "Interruptor_8" at 131,406 size 40x40

screen "Graf-cau-pot-actual" 1280x800, template "Plantilla"
   TrendView "Visor de curvas_1" at 3,109 size 1268x600
   TextField "Campo de texto_16" at 477,10 size 365x27
   TextField "Campo de texto_1" at 1143,73 size 122x25
   TextField "Campo de texto_2" at 45,70 size 137x25
   Button "Botón_1" at 271,54 size 150x40
   Button "Botón_2" at 479,54 size 150x40
   Button "Botón_3" at 687,54 size 150x40
   Button "Botón_4" at 895,54 size 150x40

screen "EcalarSeñAnal" 1280x800, template "Plantilla"
   TextField "Campo de texto_1" at 69,133 size 223x27
   TextField "Campo de texto_2" at 69,375 size 236x27
   IOField "Campo ES_1" at 415,204 size 119x32
   IOField "Campo ES_2" at 415,274 size 119x32
   IOField "Campo ES_4" at 415,451 size 119x32
   IOField "Campo ES_3" at 415,522 size 119x32
   TextField "Campo de texto_3" at 234,204 size 127x27
   TextField "Campo de texto_4" at 234,274 size 118x27
   TextField "Campo de texto_5" at 234,451 size 127x27
   TextField "Campo de texto_6" at 234,522 size 118x27
   Button "Botón_3" at 788,329 size 240x49

screen "Graf-cau-pot-historico" 1280x800, template "Plantilla"
   TrendView "Visor de curvas_1" at 3,109 size 1268x600
   TextField "Campo de texto_16" at 477,10 size 334x27
   TextField "Campo de texto_2" at 29,70 size 137x25
   TextField "Campo de texto_1" at 1143,73 size 122x25
   TextField "Campo de texto_3" at 1143,73 size 122x25
*)